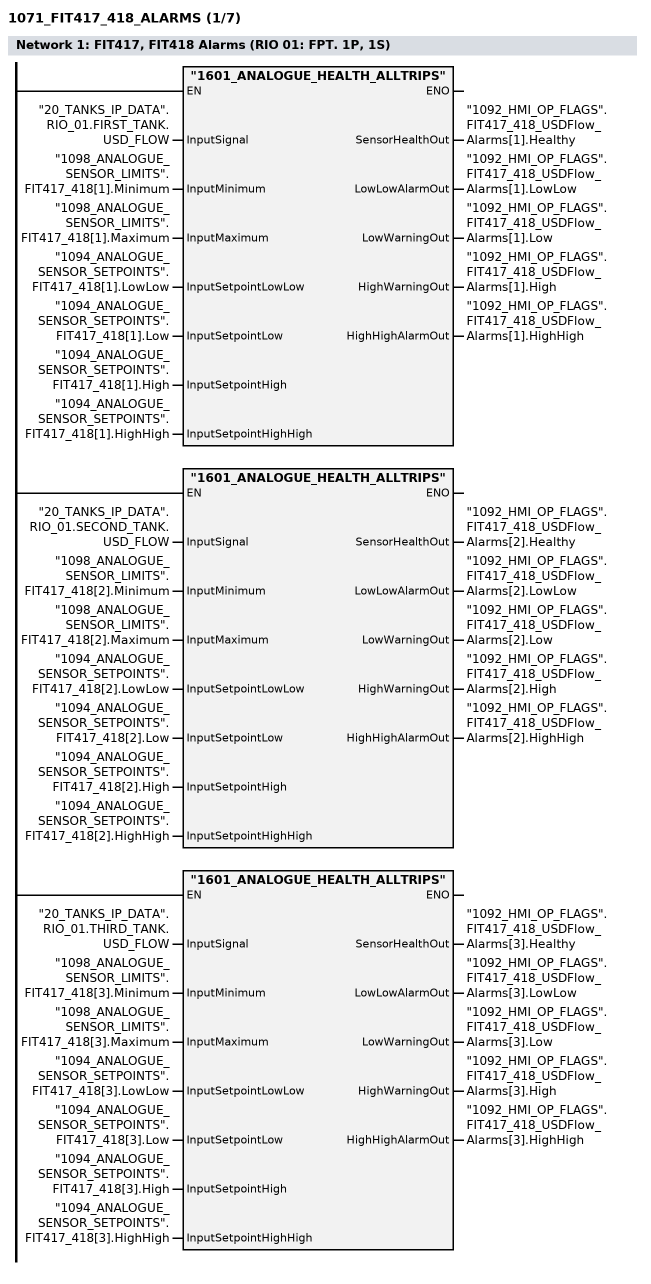
   RUNG wire#powerrail
      "1601_ANALOGUE_HEALTH_ALLTRIPS"(InputSignal := "20_TANKS_IP_DATA".RIO_01.FIRST_TANK.USD_FLOW, InputMinimum := "1098_ANALOGUE_SENSOR_LIMITS".FIT417_418[1].Minimum, InputMaximum := "1098_ANALOGUE_SENSOR_LIMITS".FIT417_418[1].Maximum, InputSetpointLowLow := "1094_ANALOGUE_SENSOR_SETPOINTS".FIT417_418[1].LowLow, InputSetpointLow := "1094_ANALOGUE_SENSOR_SETPOINTS".FIT417_418[1].Low, InputSetpointHigh := "1094_ANALOGUE_SENSOR_SETPOINTS".FIT417_418[1].High, InputSetpointHighHigh := "1094_ANALOGUE_SENSOR_SETPOINTS".FIT417_418[1].HighHigh, SensorHealthOut => "1092_HMI_OP_FLAGS".FIT417_418_USDFlow_Alarms[1].Healthy, LowLowAlarmOut => "1092_HMI_OP_FLAGS".FIT417_418_USDFlow_Alarms[1].LowLow, LowWarningOut => "1092_HMI_OP_FLAGS".FIT417_418_USDFlow_Alarms[1].Low, HighWarningOut => "1092_HMI_OP_FLAGS".FIT417_418_USDFlow_Alarms[1].High, HighHighAlarmOut => "1092_HMI_OP_FLAGS".FIT417_418_USDFlow_Alarms[1].HighHigh)
   END_RUNG
   RUNG wire#powerrail
      "1601_ANALOGUE_HEALTH_ALLTRIPS"(InputSignal := "20_TANKS_IP_DATA".RIO_01.SECOND_TANK.USD_FLOW, InputMinimum := "1098_ANALOGUE_SENSOR_LIMITS".FIT417_418[2].Minimum, InputMaximum := "1098_ANALOGUE_SENSOR_LIMITS".FIT417_418[2].Maximum, InputSetpointLowLow := "1094_ANALOGUE_SENSOR_SETPOINTS".FIT417_418[2].LowLow, InputSetpointLow := "1094_ANALOGUE_SENSOR_SETPOINTS".FIT417_418[2].Low, InputSetpointHigh := "1094_ANALOGUE_SENSOR_SETPOINTS".FIT417_418[2].High, InputSetpointHighHigh := "1094_ANALOGUE_SENSOR_SETPOINTS".FIT417_418[2].HighHigh, SensorHealthOut => "1092_HMI_OP_FLAGS".FIT417_418_USDFlow_Alarms[2].Healthy, LowLowAlarmOut => "1092_HMI_OP_FLAGS".FIT417_418_USDFlow_Alarms[2].LowLow, LowWarningOut => "1092_HMI_OP_FLAGS".FIT417_418_USDFlow_Alarms[2].Low, HighWarningOut => "1092_HMI_OP_FLAGS".FIT417_418_USDFlow_Alarms[2].High, HighHighAlarmOut => "1092_HMI_OP_FLAGS".FIT417_418_USDFlow_Alarms[2].HighHigh)
   END_RUNG
   RUNG wire#powerrail
      "1601_ANALOGUE_HEALTH_ALLTRIPS"(InputSignal := "20_TANKS_IP_DATA".RIO_01.THIRD_TANK.USD_FLOW, InputMinimum := "1098_ANALOGUE_SENSOR_LIMITS".FIT417_418[3].Minimum, InputMaximum := "1098_ANALOGUE_SENSOR_LIMITS".FIT417_418[3].Maximum, InputSetpointLowLow := "1094_ANALOGUE_SENSOR_SETPOINTS".FIT417_418[3].LowLow, InputSetpointLow := "1094_ANALOGUE_SENSOR_SETPOINTS".FIT417_418[3].Low, InputSetpointHigh := "1094_ANALOGUE_SENSOR_SETPOINTS".FIT417_418[3].High, InputSetpointHighHigh := "1094_ANALOGUE_SENSOR_SETPOINTS".FIT417_418[3].HighHigh, SensorHealthOut => "1092_HMI_OP_FLAGS".FIT417_418_USDFlow_Alarms[3].Healthy, LowLowAlarmOut => "1092_HMI_OP_FLAGS".FIT417_418_USDFlow_Alarms[3].LowLow, LowWarningOut => "1092_HMI_OP_FLAGS".FIT417_418_USDFlow_Alarms[3].Low, HighWarningOut => "1092_HMI_OP_FLAGS".FIT417_418_USDFlow_Alarms[3].High, HighHighAlarmOut => "1092_HMI_OP_FLAGS".FIT417_418_USDFlow_Alarms[3].HighHigh)
   END_RUNG
   // the same network as SCL:
   "1601_ANALOGUE_HEALTH_ALLTRIPS"(InputSignal := "20_TANKS_IP_DATA".RIO_01.FIRST_TANK.USD_FLOW,
                           InputMinimum := "1098_ANALOGUE_SENSOR_LIMITS".FIT417_418[1].Minimum,
                           InputMaximum := "1098_ANALOGUE_SENSOR_LIMITS".FIT417_418[1].Maximum,
                           InputSetpointLowLow := "1094_ANALOGUE_SENSOR_SETPOINTS".FIT417_418[1].LowLow,
                           InputSetpointLow := "1094_ANALOGUE_SENSOR_SETPOINTS".FIT417_418[1].Low,
                           InputSetpointHigh := "1094_ANALOGUE_SENSOR_SETPOINTS".FIT417_418[1].High,
                           InputSetpointHighHigh := "1094_ANALOGUE_SENSOR_SETPOINTS".FIT417_418[1].HighHigh,
                           SensorHealthOut => "1092_HMI_OP_FLAGS".FIT417_418_USDFlow_Alarms[1].Healthy,
                           LowLowAlarmOut => "1092_HMI_OP_FLAGS".FIT417_418_USDFlow_Alarms[1].LowLow,
                           LowWarningOut => "1092_HMI_OP_FLAGS".FIT417_418_USDFlow_Alarms[1].Low,
                           HighWarningOut => "1092_HMI_OP_FLAGS".FIT417_418_USDFlow_Alarms[1].High,
                           HighHighAlarmOut => "1092_HMI_OP_FLAGS".FIT417_418_USDFlow_Alarms[1].HighHigh);
   "1601_ANALOGUE_HEALTH_ALLTRIPS"(InputSignal := "20_TANKS_IP_DATA".RIO_01.SECOND_TANK.USD_FLOW,
                           InputMinimum := "1098_ANALOGUE_SENSOR_LIMITS".FIT417_418[2].Minimum,
                           InputMaximum := "1098_ANALOGUE_SENSOR_LIMITS".FIT417_418[2].Maximum,
                           InputSetpointLowLow := "1094_ANALOGUE_SENSOR_SETPOINTS".FIT417_418[2].LowLow,
                           InputSetpointLow := "1094_ANALOGUE_SENSOR_SETPOINTS".FIT417_418[2].Low,
                           InputSetpointHigh := "1094_ANALOGUE_SENSOR_SETPOINTS".FIT417_418[2].High,
                           InputSetpointHighHigh := "1094_ANALOGUE_SENSOR_SETPOINTS".FIT417_418[2].HighHigh,
                           SensorHealthOut => "1092_HMI_OP_FLAGS".FIT417_418_USDFlow_Alarms[2].Healthy,
                           LowLowAlarmOut => "1092_HMI_OP_FLAGS".FIT417_418_USDFlow_Alarms[2].LowLow,
                           LowWarningOut => "1092_HMI_OP_FLAGS".FIT417_418_USDFlow_Alarms[2].Low,
                           HighWarningOut => "1092_HMI_OP_FLAGS".FIT417_418_USDFlow_Alarms[2].High,
                           HighHighAlarmOut => "1092_HMI_OP_FLAGS".FIT417_418_USDFlow_Alarms[2].HighHigh);
   "1601_ANALOGUE_HEALTH_ALLTRIPS"(InputSignal := "20_TANKS_IP_DATA".RIO_01.THIRD_TANK.USD_FLOW,
                           InputMinimum := "1098_ANALOGUE_SENSOR_LIMITS".FIT417_418[3].Minimum,
                           InputMaximum := "1098_ANALOGUE_SENSOR_LIMITS".FIT417_418[3].Maximum,
                           InputSetpointLowLow := "1094_ANALOGUE_SENSOR_SETPOINTS".FIT417_418[3].LowLow,
                           InputSetpointLow := "1094_ANALOGUE_SENSOR_SETPOINTS".FIT417_418[3].Low,
                           InputSetpointHigh := "1094_ANALOGUE_SENSOR_SETPOINTS".FIT417_418[3].High,
                           InputSetpointHighHigh := "1094_ANALOGUE_SENSOR_SETPOINTS".FIT417_418[3].HighHigh,
                           SensorHealthOut => "1092_HMI_OP_FLAGS".FIT417_418_USDFlow_Alarms[3].Healthy,
                           LowLowAlarmOut => "1092_HMI_OP_FLAGS".FIT417_418_USDFlow_Alarms[3].LowLow,
                           LowWarningOut => "1092_HMI_OP_FLAGS".FIT417_418_USDFlow_Alarms[3].Low,
                           HighWarningOut => "1092_HMI_OP_FLAGS".FIT417_418_USDFlow_Alarms[3].High,
                           HighHighAlarmOut => "1092_HMI_OP_FLAGS".FIT417_418_USDFlow_Alarms[3].HighHigh);
END_REGION

REGION Network 2: FIT417, FIT418 Alarms (RIO 02: 2P, 2S)
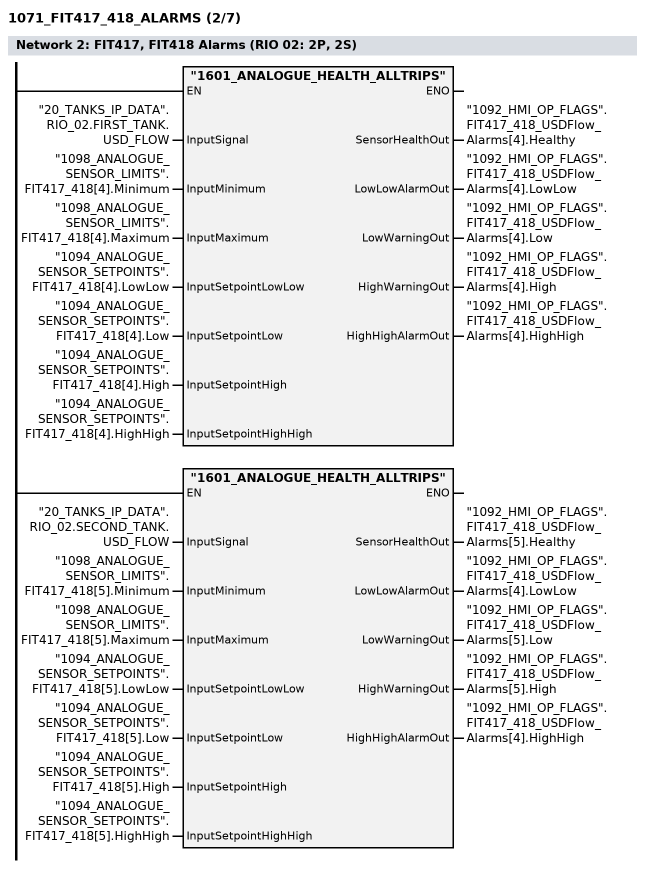
   RUNG wire#powerrail
      "1601_ANALOGUE_HEALTH_ALLTRIPS"(InputSignal := "20_TANKS_IP_DATA".RIO_02.FIRST_TANK.USD_FLOW, InputMinimum := "1098_ANALOGUE_SENSOR_LIMITS".FIT417_418[4].Minimum, InputMaximum := "1098_ANALOGUE_SENSOR_LIMITS".FIT417_418[4].Maximum, InputSetpointLowLow := "1094_ANALOGUE_SENSOR_SETPOINTS".FIT417_418[4].LowLow, InputSetpointLow := "1094_ANALOGUE_SENSOR_SETPOINTS".FIT417_418[4].Low, InputSetpointHigh := "1094_ANALOGUE_SENSOR_SETPOINTS".FIT417_418[4].High, InputSetpointHighHigh := "1094_ANALOGUE_SENSOR_SETPOINTS".FIT417_418[4].HighHigh, SensorHealthOut => "1092_HMI_OP_FLAGS".FIT417_418_USDFlow_Alarms[4].Healthy, LowLowAlarmOut => "1092_HMI_OP_FLAGS".FIT417_418_USDFlow_Alarms[4].LowLow, LowWarningOut => "1092_HMI_OP_FLAGS".FIT417_418_USDFlow_Alarms[4].Low, HighWarningOut => "1092_HMI_OP_FLAGS".FIT417_418_USDFlow_Alarms[4].High, HighHighAlarmOut => "1092_HMI_OP_FLAGS".FIT417_418_USDFlow_Alarms[4].HighHigh)
   END_RUNG
   RUNG wire#powerrail
      "1601_ANALOGUE_HEALTH_ALLTRIPS"(InputSignal := "20_TANKS_IP_DATA".RIO_02.SECOND_TANK.USD_FLOW, InputMinimum := "1098_ANALOGUE_SENSOR_LIMITS".FIT417_418[5].Minimum, InputMaximum := "1098_ANALOGUE_SENSOR_LIMITS".FIT417_418[5].Maximum, InputSetpointLowLow := "1094_ANALOGUE_SENSOR_SETPOINTS".FIT417_418[5].LowLow, InputSetpointLow := "1094_ANALOGUE_SENSOR_SETPOINTS".FIT417_418[5].Low, InputSetpointHigh := "1094_ANALOGUE_SENSOR_SETPOINTS".FIT417_418[5].High, InputSetpointHighHigh := "1094_ANALOGUE_SENSOR_SETPOINTS".FIT417_418[5].HighHigh, SensorHealthOut => "1092_HMI_OP_FLAGS".FIT417_418_USDFlow_Alarms[5].Healthy, LowLowAlarmOut => "1092_HMI_OP_FLAGS".FIT417_418_USDFlow_Alarms[4].LowLow, LowWarningOut => "1092_HMI_OP_FLAGS".FIT417_418_USDFlow_Alarms[5].Low, HighWarningOut => "1092_HMI_OP_FLAGS".FIT417_418_USDFlow_Alarms[5].High, HighHighAlarmOut => "1092_HMI_OP_FLAGS".FIT417_418_USDFlow_Alarms[4].HighHigh)
   END_RUNG
   // the same network as SCL:
   "1601_ANALOGUE_HEALTH_ALLTRIPS"(InputSignal := "20_TANKS_IP_DATA".RIO_02.FIRST_TANK.USD_FLOW,
                           InputMinimum := "1098_ANALOGUE_SENSOR_LIMITS".FIT417_418[4].Minimum,
                           InputMaximum := "1098_ANALOGUE_SENSOR_LIMITS".FIT417_418[4].Maximum,
                           InputSetpointLowLow := "1094_ANALOGUE_SENSOR_SETPOINTS".FIT417_418[4].LowLow,
                           InputSetpointLow := "1094_ANALOGUE_SENSOR_SETPOINTS".FIT417_418[4].Low,
                           InputSetpointHigh := "1094_ANALOGUE_SENSOR_SETPOINTS".FIT417_418[4].High,
                           InputSetpointHighHigh := "1094_ANALOGUE_SENSOR_SETPOINTS".FIT417_418[4].HighHigh,
                           SensorHealthOut => "1092_HMI_OP_FLAGS".FIT417_418_USDFlow_Alarms[4].Healthy,
                           LowLowAlarmOut => "1092_HMI_OP_FLAGS".FIT417_418_USDFlow_Alarms[4].LowLow,
                           LowWarningOut => "1092_HMI_OP_FLAGS".FIT417_418_USDFlow_Alarms[4].Low,
                           HighWarningOut => "1092_HMI_OP_FLAGS".FIT417_418_USDFlow_Alarms[4].High,
                           HighHighAlarmOut => "1092_HMI_OP_FLAGS".FIT417_418_USDFlow_Alarms[4].HighHigh);
   "1601_ANALOGUE_HEALTH_ALLTRIPS"(InputSignal := "20_TANKS_IP_DATA".RIO_02.SECOND_TANK.USD_FLOW,
                           InputMinimum := "1098_ANALOGUE_SENSOR_LIMITS".FIT417_418[5].Minimum,
                           InputMaximum := "1098_ANALOGUE_SENSOR_LIMITS".FIT417_418[5].Maximum,
                           InputSetpointLowLow := "1094_ANALOGUE_SENSOR_SETPOINTS".FIT417_418[5].LowLow,
                           InputSetpointLow := "1094_ANALOGUE_SENSOR_SETPOINTS".FIT417_418[5].Low,
                           InputSetpointHigh := "1094_ANALOGUE_SENSOR_SETPOINTS".FIT417_418[5].High,
                           InputSetpointHighHigh := "1094_ANALOGUE_SENSOR_SETPOINTS".FIT417_418[5].HighHigh,
                           SensorHealthOut => "1092_HMI_OP_FLAGS".FIT417_418_USDFlow_Alarms[5].Healthy,
                           LowLowAlarmOut => "1092_HMI_OP_FLAGS".FIT417_418_USDFlow_Alarms[4].LowLow,
                           LowWarningOut => "1092_HMI_OP_FLAGS".FIT417_418_USDFlow_Alarms[5].Low,
                           HighWarningOut => "1092_HMI_OP_FLAGS".FIT417_418_USDFlow_Alarms[5].High,
                           HighHighAlarmOut => "1092_HMI_OP_FLAGS".FIT417_418_USDFlow_Alarms[4].HighHigh);
END_REGION

REGION Network 3: FIT417, FIT418 Alarms (RIO 03: 3P, 3S)
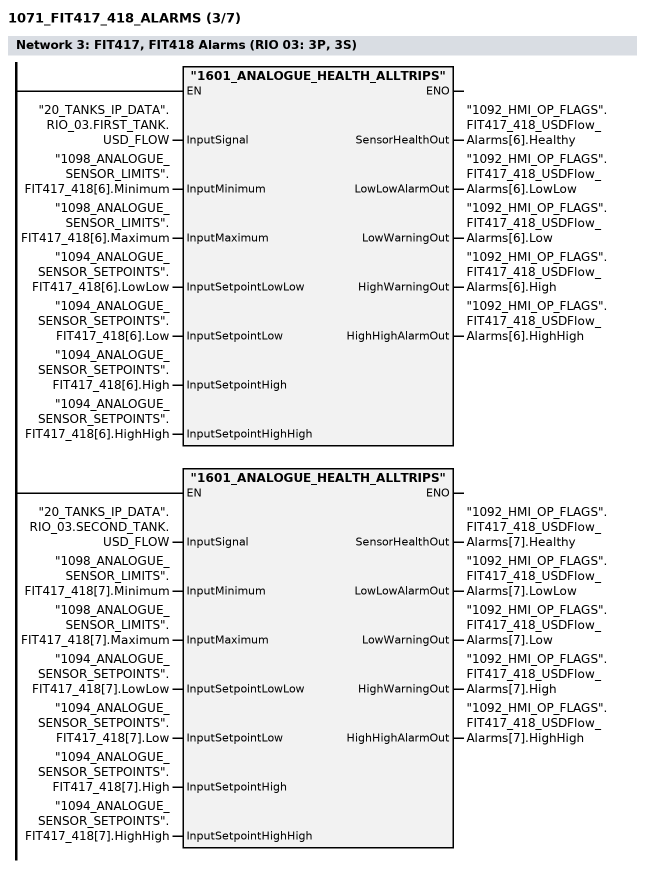
   RUNG wire#powerrail
      "1601_ANALOGUE_HEALTH_ALLTRIPS"(InputSignal := "20_TANKS_IP_DATA".RIO_03.FIRST_TANK.USD_FLOW, InputMinimum := "1098_ANALOGUE_SENSOR_LIMITS".FIT417_418[6].Minimum, InputMaximum := "1098_ANALOGUE_SENSOR_LIMITS".FIT417_418[6].Maximum, InputSetpointLowLow := "1094_ANALOGUE_SENSOR_SETPOINTS".FIT417_418[6].LowLow, InputSetpointLow := "1094_ANALOGUE_SENSOR_SETPOINTS".FIT417_418[6].Low, InputSetpointHigh := "1094_ANALOGUE_SENSOR_SETPOINTS".FIT417_418[6].High, InputSetpointHighHigh := "1094_ANALOGUE_SENSOR_SETPOINTS".FIT417_418[6].HighHigh, SensorHealthOut => "1092_HMI_OP_FLAGS".FIT417_418_USDFlow_Alarms[6].Healthy, LowLowAlarmOut => "1092_HMI_OP_FLAGS".FIT417_418_USDFlow_Alarms[6].LowLow, LowWarningOut => "1092_HMI_OP_FLAGS".FIT417_418_USDFlow_Alarms[6].Low, HighWarningOut => "1092_HMI_OP_FLAGS".FIT417_418_USDFlow_Alarms[6].High, HighHighAlarmOut => "1092_HMI_OP_FLAGS".FIT417_418_USDFlow_Alarms[6].HighHigh)
   END_RUNG
   RUNG wire#powerrail
      "1601_ANALOGUE_HEALTH_ALLTRIPS"(InputSignal := "20_TANKS_IP_DATA".RIO_03.SECOND_TANK.USD_FLOW, InputMinimum := "1098_ANALOGUE_SENSOR_LIMITS".FIT417_418[7].Minimum, InputMaximum := "1098_ANALOGUE_SENSOR_LIMITS".FIT417_418[7].Maximum, InputSetpointLowLow := "1094_ANALOGUE_SENSOR_SETPOINTS".FIT417_418[7].LowLow, InputSetpointLow := "1094_ANALOGUE_SENSOR_SETPOINTS".FIT417_418[7].Low, InputSetpointHigh := "1094_ANALOGUE_SENSOR_SETPOINTS".FIT417_418[7].High, InputSetpointHighHigh := "1094_ANALOGUE_SENSOR_SETPOINTS".FIT417_418[7].HighHigh, SensorHealthOut => "1092_HMI_OP_FLAGS".FIT417_418_USDFlow_Alarms[7].Healthy, LowLowAlarmOut => "1092_HMI_OP_FLAGS".FIT417_418_USDFlow_Alarms[7].LowLow, LowWarningOut => "1092_HMI_OP_FLAGS".FIT417_418_USDFlow_Alarms[7].Low, HighWarningOut => "1092_HMI_OP_FLAGS".FIT417_418_USDFlow_Alarms[7].High, HighHighAlarmOut => "1092_HMI_OP_FLAGS".FIT417_418_USDFlow_Alarms[7].HighHigh)
   END_RUNG
   // the same network as SCL:
   "1601_ANALOGUE_HEALTH_ALLTRIPS"(InputSignal := "20_TANKS_IP_DATA".RIO_03.FIRST_TANK.USD_FLOW,
                           InputMinimum := "1098_ANALOGUE_SENSOR_LIMITS".FIT417_418[6].Minimum,
                           InputMaximum := "1098_ANALOGUE_SENSOR_LIMITS".FIT417_418[6].Maximum,
                           InputSetpointLowLow := "1094_ANALOGUE_SENSOR_SETPOINTS".FIT417_418[6].LowLow,
                           InputSetpointLow := "1094_ANALOGUE_SENSOR_SETPOINTS".FIT417_418[6].Low,
                           InputSetpointHigh := "1094_ANALOGUE_SENSOR_SETPOINTS".FIT417_418[6].High,
                           InputSetpointHighHigh := "1094_ANALOGUE_SENSOR_SETPOINTS".FIT417_418[6].HighHigh,
                           SensorHealthOut => "1092_HMI_OP_FLAGS".FIT417_418_USDFlow_Alarms[6].Healthy,
                           LowLowAlarmOut => "1092_HMI_OP_FLAGS".FIT417_418_USDFlow_Alarms[6].LowLow,
                           LowWarningOut => "1092_HMI_OP_FLAGS".FIT417_418_USDFlow_Alarms[6].Low,
                           HighWarningOut => "1092_HMI_OP_FLAGS".FIT417_418_USDFlow_Alarms[6].High,
                           HighHighAlarmOut => "1092_HMI_OP_FLAGS".FIT417_418_USDFlow_Alarms[6].HighHigh);
   "1601_ANALOGUE_HEALTH_ALLTRIPS"(InputSignal := "20_TANKS_IP_DATA".RIO_03.SECOND_TANK.USD_FLOW,
                           InputMinimum := "1098_ANALOGUE_SENSOR_LIMITS".FIT417_418[7].Minimum,
                           InputMaximum := "1098_ANALOGUE_SENSOR_LIMITS".FIT417_418[7].Maximum,
                           InputSetpointLowLow := "1094_ANALOGUE_SENSOR_SETPOINTS".FIT417_418[7].LowLow,
                           InputSetpointLow := "1094_ANALOGUE_SENSOR_SETPOINTS".FIT417_418[7].Low,
                           InputSetpointHigh := "1094_ANALOGUE_SENSOR_SETPOINTS".FIT417_418[7].High,
                           InputSetpointHighHigh := "1094_ANALOGUE_SENSOR_SETPOINTS".FIT417_418[7].HighHigh,
                           SensorHealthOut => "1092_HMI_OP_FLAGS".FIT417_418_USDFlow_Alarms[7].Healthy,
                           LowLowAlarmOut => "1092_HMI_OP_FLAGS".FIT417_418_USDFlow_Alarms[7].LowLow,
                           LowWarningOut => "1092_HMI_OP_FLAGS".FIT417_418_USDFlow_Alarms[7].Low,
                           HighWarningOut => "1092_HMI_OP_FLAGS".FIT417_418_USDFlow_Alarms[7].High,
                           HighHighAlarmOut => "1092_HMI_OP_FLAGS".FIT417_418_USDFlow_Alarms[7].HighHigh);
END_REGION

REGION Network 4: FIT417, FIT418 Alarms (RIO 04: 4P, 4S)
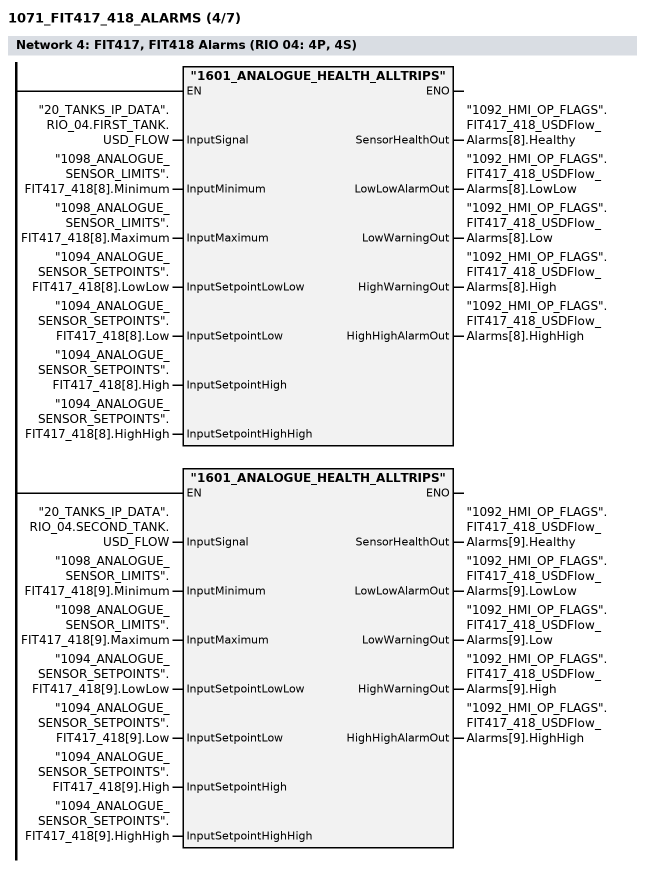
   RUNG wire#powerrail
      "1601_ANALOGUE_HEALTH_ALLTRIPS"(InputSignal := "20_TANKS_IP_DATA".RIO_04.FIRST_TANK.USD_FLOW, InputMinimum := "1098_ANALOGUE_SENSOR_LIMITS".FIT417_418[8].Minimum, InputMaximum := "1098_ANALOGUE_SENSOR_LIMITS".FIT417_418[8].Maximum, InputSetpointLowLow := "1094_ANALOGUE_SENSOR_SETPOINTS".FIT417_418[8].LowLow, InputSetpointLow := "1094_ANALOGUE_SENSOR_SETPOINTS".FIT417_418[8].Low, InputSetpointHigh := "1094_ANALOGUE_SENSOR_SETPOINTS".FIT417_418[8].High, InputSetpointHighHigh := "1094_ANALOGUE_SENSOR_SETPOINTS".FIT417_418[8].HighHigh, SensorHealthOut => "1092_HMI_OP_FLAGS".FIT417_418_USDFlow_Alarms[8].Healthy, LowLowAlarmOut => "1092_HMI_OP_FLAGS".FIT417_418_USDFlow_Alarms[8].LowLow, LowWarningOut => "1092_HMI_OP_FLAGS".FIT417_418_USDFlow_Alarms[8].Low, HighWarningOut => "1092_HMI_OP_FLAGS".FIT417_418_USDFlow_Alarms[8].High, HighHighAlarmOut => "1092_HMI_OP_FLAGS".FIT417_418_USDFlow_Alarms[8].HighHigh)
   END_RUNG
   RUNG wire#powerrail
      "1601_ANALOGUE_HEALTH_ALLTRIPS"(InputSignal := "20_TANKS_IP_DATA".RIO_04.SECOND_TANK.USD_FLOW, InputMinimum := "1098_ANALOGUE_SENSOR_LIMITS".FIT417_418[9].Minimum, InputMaximum := "1098_ANALOGUE_SENSOR_LIMITS".FIT417_418[9].Maximum, InputSetpointLowLow := "1094_ANALOGUE_SENSOR_SETPOINTS".FIT417_418[9].LowLow, InputSetpointLow := "1094_ANALOGUE_SENSOR_SETPOINTS".FIT417_418[9].Low, InputSetpointHigh := "1094_ANALOGUE_SENSOR_SETPOINTS".FIT417_418[9].High, InputSetpointHighHigh := "1094_ANALOGUE_SENSOR_SETPOINTS".FIT417_418[9].HighHigh, SensorHealthOut => "1092_HMI_OP_FLAGS".FIT417_418_USDFlow_Alarms[9].Healthy, LowLowAlarmOut => "1092_HMI_OP_FLAGS".FIT417_418_USDFlow_Alarms[9].LowLow, LowWarningOut => "1092_HMI_OP_FLAGS".FIT417_418_USDFlow_Alarms[9].Low, HighWarningOut => "1092_HMI_OP_FLAGS".FIT417_418_USDFlow_Alarms[9].High, HighHighAlarmOut => "1092_HMI_OP_FLAGS".FIT417_418_USDFlow_Alarms[9].HighHigh)
   END_RUNG
   // the same network as SCL:
   "1601_ANALOGUE_HEALTH_ALLTRIPS"(InputSignal := "20_TANKS_IP_DATA".RIO_04.FIRST_TANK.USD_FLOW,
                           InputMinimum := "1098_ANALOGUE_SENSOR_LIMITS".FIT417_418[8].Minimum,
                           InputMaximum := "1098_ANALOGUE_SENSOR_LIMITS".FIT417_418[8].Maximum,
                           InputSetpointLowLow := "1094_ANALOGUE_SENSOR_SETPOINTS".FIT417_418[8].LowLow,
                           InputSetpointLow := "1094_ANALOGUE_SENSOR_SETPOINTS".FIT417_418[8].Low,
                           InputSetpointHigh := "1094_ANALOGUE_SENSOR_SETPOINTS".FIT417_418[8].High,
                           InputSetpointHighHigh := "1094_ANALOGUE_SENSOR_SETPOINTS".FIT417_418[8].HighHigh,
                           SensorHealthOut => "1092_HMI_OP_FLAGS".FIT417_418_USDFlow_Alarms[8].Healthy,
                           LowLowAlarmOut => "1092_HMI_OP_FLAGS".FIT417_418_USDFlow_Alarms[8].LowLow,
                           LowWarningOut => "1092_HMI_OP_FLAGS".FIT417_418_USDFlow_Alarms[8].Low,
                           HighWarningOut => "1092_HMI_OP_FLAGS".FIT417_418_USDFlow_Alarms[8].High,
                           HighHighAlarmOut => "1092_HMI_OP_FLAGS".FIT417_418_USDFlow_Alarms[8].HighHigh);
   "1601_ANALOGUE_HEALTH_ALLTRIPS"(InputSignal := "20_TANKS_IP_DATA".RIO_04.SECOND_TANK.USD_FLOW,
                           InputMinimum := "1098_ANALOGUE_SENSOR_LIMITS".FIT417_418[9].Minimum,
                           InputMaximum := "1098_ANALOGUE_SENSOR_LIMITS".FIT417_418[9].Maximum,
                           InputSetpointLowLow := "1094_ANALOGUE_SENSOR_SETPOINTS".FIT417_418[9].LowLow,
                           InputSetpointLow := "1094_ANALOGUE_SENSOR_SETPOINTS".FIT417_418[9].Low,
                           InputSetpointHigh := "1094_ANALOGUE_SENSOR_SETPOINTS".FIT417_418[9].High,
                           InputSetpointHighHigh := "1094_ANALOGUE_SENSOR_SETPOINTS".FIT417_418[9].HighHigh,
                           SensorHealthOut => "1092_HMI_OP_FLAGS".FIT417_418_USDFlow_Alarms[9].Healthy,
                           LowLowAlarmOut => "1092_HMI_OP_FLAGS".FIT417_418_USDFlow_Alarms[9].LowLow,
                           LowWarningOut => "1092_HMI_OP_FLAGS".FIT417_418_USDFlow_Alarms[9].Low,
                           HighWarningOut => "1092_HMI_OP_FLAGS".FIT417_418_USDFlow_Alarms[9].High,
                           HighHighAlarmOut => "1092_HMI_OP_FLAGS".FIT417_418_USDFlow_Alarms[9].HighHigh);
END_REGION

REGION Network 5: FIT417, FIT418 Alarms (RIO 05: 5P, 5S)
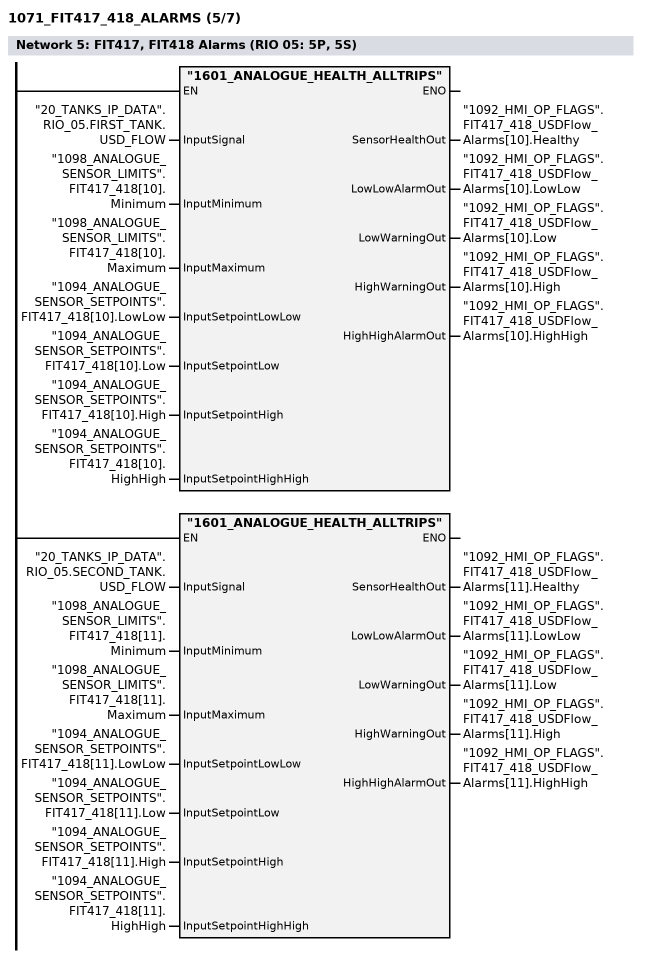
   RUNG wire#powerrail
      "1601_ANALOGUE_HEALTH_ALLTRIPS"(InputSignal := "20_TANKS_IP_DATA".RIO_05.FIRST_TANK.USD_FLOW, InputMinimum := "1098_ANALOGUE_SENSOR_LIMITS".FIT417_418[10].Minimum, InputMaximum := "1098_ANALOGUE_SENSOR_LIMITS".FIT417_418[10].Maximum, InputSetpointLowLow := "1094_ANALOGUE_SENSOR_SETPOINTS".FIT417_418[10].LowLow, InputSetpointLow := "1094_ANALOGUE_SENSOR_SETPOINTS".FIT417_418[10].Low, InputSetpointHigh := "1094_ANALOGUE_SENSOR_SETPOINTS".FIT417_418[10].High, InputSetpointHighHigh := "1094_ANALOGUE_SENSOR_SETPOINTS".FIT417_418[10].HighHigh, SensorHealthOut => "1092_HMI_OP_FLAGS".FIT417_418_USDFlow_Alarms[10].Healthy, LowLowAlarmOut => "1092_HMI_OP_FLAGS".FIT417_418_USDFlow_Alarms[10].LowLow, LowWarningOut => "1092_HMI_OP_FLAGS".FIT417_418_USDFlow_Alarms[10].Low, HighWarningOut => "1092_HMI_OP_FLAGS".FIT417_418_USDFlow_Alarms[10].High, HighHighAlarmOut => "1092_HMI_OP_FLAGS".FIT417_418_USDFlow_Alarms[10].HighHigh)
   END_RUNG
   RUNG wire#powerrail
      "1601_ANALOGUE_HEALTH_ALLTRIPS"(InputSignal := "20_TANKS_IP_DATA".RIO_05.SECOND_TANK.USD_FLOW, InputMinimum := "1098_ANALOGUE_SENSOR_LIMITS".FIT417_418[11].Minimum, InputMaximum := "1098_ANALOGUE_SENSOR_LIMITS".FIT417_418[11].Maximum, InputSetpointLowLow := "1094_ANALOGUE_SENSOR_SETPOINTS".FIT417_418[11].LowLow, InputSetpointLow := "1094_ANALOGUE_SENSOR_SETPOINTS".FIT417_418[11].Low, InputSetpointHigh := "1094_ANALOGUE_SENSOR_SETPOINTS".FIT417_418[11].High, InputSetpointHighHigh := "1094_ANALOGUE_SENSOR_SETPOINTS".FIT417_418[11].HighHigh, SensorHealthOut => "1092_HMI_OP_FLAGS".FIT417_418_USDFlow_Alarms[11].Healthy, LowLowAlarmOut => "1092_HMI_OP_FLAGS".FIT417_418_USDFlow_Alarms[11].LowLow, LowWarningOut => "1092_HMI_OP_FLAGS".FIT417_418_USDFlow_Alarms[11].Low, HighWarningOut => "1092_HMI_OP_FLAGS".FIT417_418_USDFlow_Alarms[11].High, HighHighAlarmOut => "1092_HMI_OP_FLAGS".FIT417_418_USDFlow_Alarms[11].HighHigh)
   END_RUNG
   // the same network as SCL:
   "1601_ANALOGUE_HEALTH_ALLTRIPS"(InputSignal := "20_TANKS_IP_DATA".RIO_05.FIRST_TANK.USD_FLOW,
                           InputMinimum := "1098_ANALOGUE_SENSOR_LIMITS".FIT417_418[10].Minimum,
                           InputMaximum := "1098_ANALOGUE_SENSOR_LIMITS".FIT417_418[10].Maximum,
                           InputSetpointLowLow := "1094_ANALOGUE_SENSOR_SETPOINTS".FIT417_418[10].LowLow,
                           InputSetpointLow := "1094_ANALOGUE_SENSOR_SETPOINTS".FIT417_418[10].Low,
                           InputSetpointHigh := "1094_ANALOGUE_SENSOR_SETPOINTS".FIT417_418[10].High,
                           InputSetpointHighHigh := "1094_ANALOGUE_SENSOR_SETPOINTS".FIT417_418[10].HighHigh,
                           SensorHealthOut => "1092_HMI_OP_FLAGS".FIT417_418_USDFlow_Alarms[10].Healthy,
                           LowLowAlarmOut => "1092_HMI_OP_FLAGS".FIT417_418_USDFlow_Alarms[10].LowLow,
                           LowWarningOut => "1092_HMI_OP_FLAGS".FIT417_418_USDFlow_Alarms[10].Low,
                           HighWarningOut => "1092_HMI_OP_FLAGS".FIT417_418_USDFlow_Alarms[10].High,
                           HighHighAlarmOut => "1092_HMI_OP_FLAGS".FIT417_418_USDFlow_Alarms[10].HighHigh);
   "1601_ANALOGUE_HEALTH_ALLTRIPS"(InputSignal := "20_TANKS_IP_DATA".RIO_05.SECOND_TANK.USD_FLOW,
                           InputMinimum := "1098_ANALOGUE_SENSOR_LIMITS".FIT417_418[11].Minimum,
                           InputMaximum := "1098_ANALOGUE_SENSOR_LIMITS".FIT417_418[11].Maximum,
                           InputSetpointLowLow := "1094_ANALOGUE_SENSOR_SETPOINTS".FIT417_418[11].LowLow,
                           InputSetpointLow := "1094_ANALOGUE_SENSOR_SETPOINTS".FIT417_418[11].Low,
                           InputSetpointHigh := "1094_ANALOGUE_SENSOR_SETPOINTS".FIT417_418[11].High,
                           InputSetpointHighHigh := "1094_ANALOGUE_SENSOR_SETPOINTS".FIT417_418[11].HighHigh,
                           SensorHealthOut => "1092_HMI_OP_FLAGS".FIT417_418_USDFlow_Alarms[11].Healthy,
                           LowLowAlarmOut => "1092_HMI_OP_FLAGS".FIT417_418_USDFlow_Alarms[11].LowLow,
                           LowWarningOut => "1092_HMI_OP_FLAGS".FIT417_418_USDFlow_Alarms[11].Low,
                           HighWarningOut => "1092_HMI_OP_FLAGS".FIT417_418_USDFlow_Alarms[11].High,
                           HighHighAlarmOut => "1092_HMI_OP_FLAGS".FIT417_418_USDFlow_Alarms[11].HighHigh);
END_REGION

REGION Network 6: FIT417, FIT418 Alarms (RIO 06: 6P, 6S)
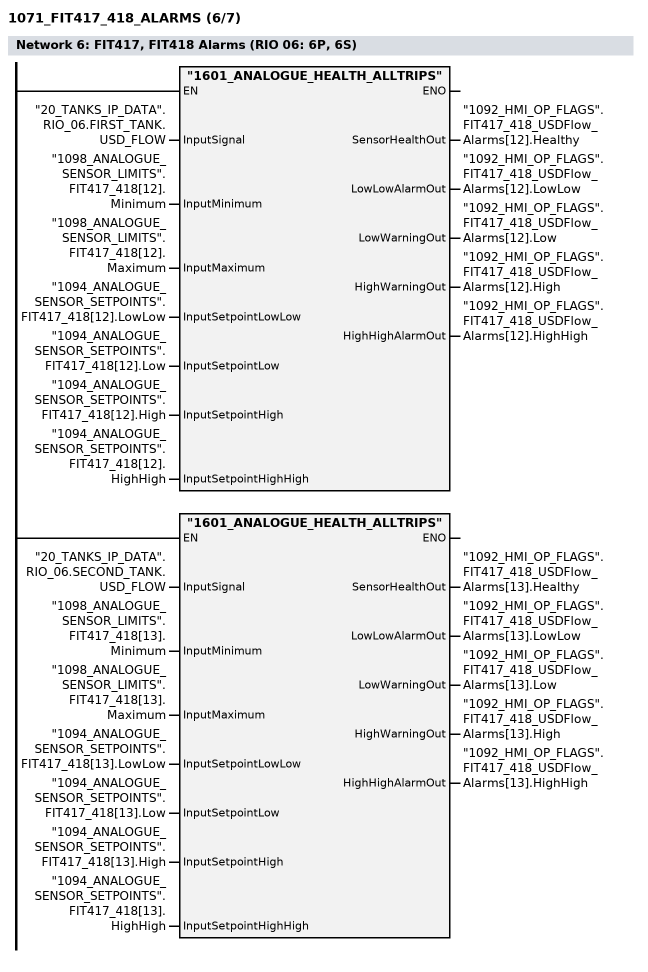
   RUNG wire#powerrail
      "1601_ANALOGUE_HEALTH_ALLTRIPS"(InputSignal := "20_TANKS_IP_DATA".RIO_06.FIRST_TANK.USD_FLOW, InputMinimum := "1098_ANALOGUE_SENSOR_LIMITS".FIT417_418[12].Minimum, InputMaximum := "1098_ANALOGUE_SENSOR_LIMITS".FIT417_418[12].Maximum, InputSetpointLowLow := "1094_ANALOGUE_SENSOR_SETPOINTS".FIT417_418[12].LowLow, InputSetpointLow := "1094_ANALOGUE_SENSOR_SETPOINTS".FIT417_418[12].Low, InputSetpointHigh := "1094_ANALOGUE_SENSOR_SETPOINTS".FIT417_418[12].High, InputSetpointHighHigh := "1094_ANALOGUE_SENSOR_SETPOINTS".FIT417_418[12].HighHigh, SensorHealthOut => "1092_HMI_OP_FLAGS".FIT417_418_USDFlow_Alarms[12].Healthy, LowLowAlarmOut => "1092_HMI_OP_FLAGS".FIT417_418_USDFlow_Alarms[12].LowLow, LowWarningOut => "1092_HMI_OP_FLAGS".FIT417_418_USDFlow_Alarms[12].Low, HighWarningOut => "1092_HMI_OP_FLAGS".FIT417_418_USDFlow_Alarms[12].High, HighHighAlarmOut => "1092_HMI_OP_FLAGS".FIT417_418_USDFlow_Alarms[12].HighHigh)
   END_RUNG
   RUNG wire#powerrail
      "1601_ANALOGUE_HEALTH_ALLTRIPS"(InputSignal := "20_TANKS_IP_DATA".RIO_06.SECOND_TANK.USD_FLOW, InputMinimum := "1098_ANALOGUE_SENSOR_LIMITS".FIT417_418[13].Minimum, InputMaximum := "1098_ANALOGUE_SENSOR_LIMITS".FIT417_418[13].Maximum, InputSetpointLowLow := "1094_ANALOGUE_SENSOR_SETPOINTS".FIT417_418[13].LowLow, InputSetpointLow := "1094_ANALOGUE_SENSOR_SETPOINTS".FIT417_418[13].Low, InputSetpointHigh := "1094_ANALOGUE_SENSOR_SETPOINTS".FIT417_418[13].High, InputSetpointHighHigh := "1094_ANALOGUE_SENSOR_SETPOINTS".FIT417_418[13].HighHigh, SensorHealthOut => "1092_HMI_OP_FLAGS".FIT417_418_USDFlow_Alarms[13].Healthy, LowLowAlarmOut => "1092_HMI_OP_FLAGS".FIT417_418_USDFlow_Alarms[13].LowLow, LowWarningOut => "1092_HMI_OP_FLAGS".FIT417_418_USDFlow_Alarms[13].Low, HighWarningOut => "1092_HMI_OP_FLAGS".FIT417_418_USDFlow_Alarms[13].High, HighHighAlarmOut => "1092_HMI_OP_FLAGS".FIT417_418_USDFlow_Alarms[13].HighHigh)
   END_RUNG
   // the same network as SCL:
   "1601_ANALOGUE_HEALTH_ALLTRIPS"(InputSignal := "20_TANKS_IP_DATA".RIO_06.FIRST_TANK.USD_FLOW,
                           InputMinimum := "1098_ANALOGUE_SENSOR_LIMITS".FIT417_418[12].Minimum,
                           InputMaximum := "1098_ANALOGUE_SENSOR_LIMITS".FIT417_418[12].Maximum,
                           InputSetpointLowLow := "1094_ANALOGUE_SENSOR_SETPOINTS".FIT417_418[12].LowLow,
                           InputSetpointLow := "1094_ANALOGUE_SENSOR_SETPOINTS".FIT417_418[12].Low,
                           InputSetpointHigh := "1094_ANALOGUE_SENSOR_SETPOINTS".FIT417_418[12].High,
                           InputSetpointHighHigh := "1094_ANALOGUE_SENSOR_SETPOINTS".FIT417_418[12].HighHigh,
                           SensorHealthOut => "1092_HMI_OP_FLAGS".FIT417_418_USDFlow_Alarms[12].Healthy,
                           LowLowAlarmOut => "1092_HMI_OP_FLAGS".FIT417_418_USDFlow_Alarms[12].LowLow,
                           LowWarningOut => "1092_HMI_OP_FLAGS".FIT417_418_USDFlow_Alarms[12].Low,
                           HighWarningOut => "1092_HMI_OP_FLAGS".FIT417_418_USDFlow_Alarms[12].High,
                           HighHighAlarmOut => "1092_HMI_OP_FLAGS".FIT417_418_USDFlow_Alarms[12].HighHigh);
   "1601_ANALOGUE_HEALTH_ALLTRIPS"(InputSignal := "20_TANKS_IP_DATA".RIO_06.SECOND_TANK.USD_FLOW,
                           InputMinimum := "1098_ANALOGUE_SENSOR_LIMITS".FIT417_418[13].Minimum,
                           InputMaximum := "1098_ANALOGUE_SENSOR_LIMITS".FIT417_418[13].Maximum,
                           InputSetpointLowLow := "1094_ANALOGUE_SENSOR_SETPOINTS".FIT417_418[13].LowLow,
                           InputSetpointLow := "1094_ANALOGUE_SENSOR_SETPOINTS".FIT417_418[13].Low,
                           InputSetpointHigh := "1094_ANALOGUE_SENSOR_SETPOINTS".FIT417_418[13].High,
                           InputSetpointHighHigh := "1094_ANALOGUE_SENSOR_SETPOINTS".FIT417_418[13].HighHigh,
                           SensorHealthOut => "1092_HMI_OP_FLAGS".FIT417_418_USDFlow_Alarms[13].Healthy,
                           LowLowAlarmOut => "1092_HMI_OP_FLAGS".FIT417_418_USDFlow_Alarms[13].LowLow,
                           LowWarningOut => "1092_HMI_OP_FLAGS".FIT417_418_USDFlow_Alarms[13].Low,
                           HighWarningOut => "1092_HMI_OP_FLAGS".FIT417_418_USDFlow_Alarms[13].High,
                           HighHighAlarmOut => "1092_HMI_OP_FLAGS".FIT417_418_USDFlow_Alarms[13].HighHigh);
END_REGION

REGION Network 7: FIT417, FIT418 Alarms (RIO 07: APT)
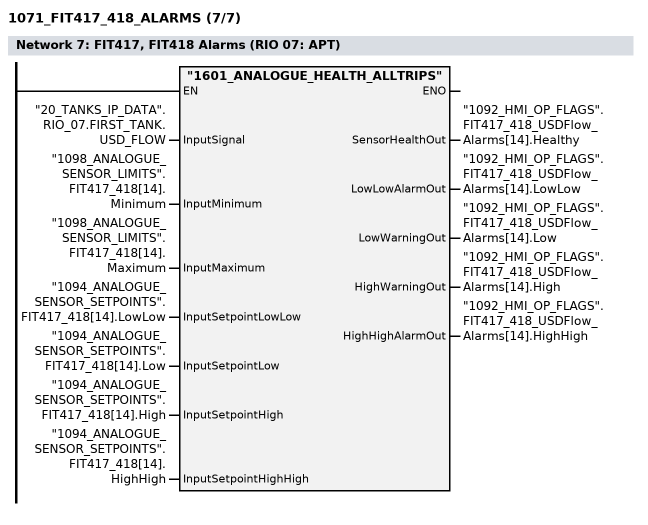
   RUNG wire#powerrail
      "1601_ANALOGUE_HEALTH_ALLTRIPS"(InputSignal := "20_TANKS_IP_DATA".RIO_07.FIRST_TANK.USD_FLOW, InputMinimum := "1098_ANALOGUE_SENSOR_LIMITS".FIT417_418[14].Minimum, InputMaximum := "1098_ANALOGUE_SENSOR_LIMITS".FIT417_418[14].Maximum, InputSetpointLowLow := "1094_ANALOGUE_SENSOR_SETPOINTS".FIT417_418[14].LowLow, InputSetpointLow := "1094_ANALOGUE_SENSOR_SETPOINTS".FIT417_418[14].Low, InputSetpointHigh := "1094_ANALOGUE_SENSOR_SETPOINTS".FIT417_418[14].High, InputSetpointHighHigh := "1094_ANALOGUE_SENSOR_SETPOINTS".FIT417_418[14].HighHigh, SensorHealthOut => "1092_HMI_OP_FLAGS".FIT417_418_USDFlow_Alarms[14].Healthy, LowLowAlarmOut => "1092_HMI_OP_FLAGS".FIT417_418_USDFlow_Alarms[14].LowLow, LowWarningOut => "1092_HMI_OP_FLAGS".FIT417_418_USDFlow_Alarms[14].Low, HighWarningOut => "1092_HMI_OP_FLAGS".FIT417_418_USDFlow_Alarms[14].High, HighHighAlarmOut => "1092_HMI_OP_FLAGS".FIT417_418_USDFlow_Alarms[14].HighHigh)
   END_RUNG
   // the same network as SCL:
   "1601_ANALOGUE_HEALTH_ALLTRIPS"(InputSignal := "20_TANKS_IP_DATA".RIO_07.FIRST_TANK.USD_FLOW,
                           InputMinimum := "1098_ANALOGUE_SENSOR_LIMITS".FIT417_418[14].Minimum,
                           InputMaximum := "1098_ANALOGUE_SENSOR_LIMITS".FIT417_418[14].Maximum,
                           InputSetpointLowLow := "1094_ANALOGUE_SENSOR_SETPOINTS".FIT417_418[14].LowLow,
                           InputSetpointLow := "1094_ANALOGUE_SENSOR_SETPOINTS".FIT417_418[14].Low,
                           InputSetpointHigh := "1094_ANALOGUE_SENSOR_SETPOINTS".FIT417_418[14].High,
                           InputSetpointHighHigh := "1094_ANALOGUE_SENSOR_SETPOINTS".FIT417_418[14].HighHigh,
                           SensorHealthOut => "1092_HMI_OP_FLAGS".FIT417_418_USDFlow_Alarms[14].Healthy,
                           LowLowAlarmOut => "1092_HMI_OP_FLAGS".FIT417_418_USDFlow_Alarms[14].LowLow,
                           LowWarningOut => "1092_HMI_OP_FLAGS".FIT417_418_USDFlow_Alarms[14].Low,
                           HighWarningOut => "1092_HMI_OP_FLAGS".FIT417_418_USDFlow_Alarms[14].High,
                           HighHighAlarmOut => "1092_HMI_OP_FLAGS".FIT417_418_USDFlow_Alarms[14].HighHigh);
END_REGION
END_FUNCTION

FUNCTION "1072_FIT419_420_ALARMS" : Void   // FC1072, LAD
{ S7_Optimized_Access := 'TRUE' }
VERSION : 0.1
// Alarm wrapper function for MBG Flow on each tank.
BEGIN

REGION Network 1: FIT419, FIT420 Alarms (RIO 01: FPT. 1P, 1S)
